// TIA Portal project "Mawomat" (V17) (continued)

               END_IF;

           ELSIF NOT #statSwitchControl OR NOT #statSwitchEnable THEN //if no output enable or switch check then

               IF #statControl THEN

                   #oStatus := 8;

               ELSIF NOT #statControl THEN

                   #oStatus := 2;

               END_IF;

           END_IF;

       ELSE
           #oStatus := 0;

       END_IF;

   END_REGION ;


   REGION Reseting impuls
       // Samokasowanie sygnalow
       #statFaultReset := false;

       IF #inAutoOff THEN

           #statTurnOn := FALSE;

       END_IF;

   END_REGION ;

   REGION Status code


   END_REGION

   REGION Rewriting TO outputs

       #inCmdOper.%X0 := #statManAuto;
       #inCmdOper.%X1 := #statSymOn;
       #inCmdOper.%X2 := #statSwitchEnable;
       #inCmdOper.%X3 := #statManTurnOn;
       #inCmdOper.%X4 := #statManDirection;
       #inCmdOper.%X6 := #statSwitchControl;

       #inCmdOperImp.%X0 := #statFaultReset;

       #oControlMode := #statControlMode;

       #oFault := #statFault;

       #inTurnOn := #statTurnOn;

       #oControl := #statControl;

   END_REGION
END_FUNCTION_BLOCK

// folder: DV

FUNCTION_BLOCK "DV_Objects"   // FB6, LAD
{ S7_Optimized_Access := 'TRUE' }
VERSION : 0.1
   VAR
      dv1 : "DV_Class";
   END_VAR
BEGIN

REGION Network 2 (SCL)
   #dv1();
END_REGION
END_FUNCTION_BLOCK

FUNCTION_BLOCK "DV_Class"   // FB302, SCL
{ S7_Optimized_Access := 'TRUE' }
VERSION : 0.1
   VAR_INPUT
      inActivateObject : Bool := true;   // Aktywowanie działania obiektu
      inTurnOnConfirm : Bool;   // Potwierdzenie załączenia
      inTurnOffConfirm : Bool;   // Potwierdzenie wyłączenia
      inCircBreaker : Bool;   // Gotowość obiektu - rozłącznik
      inPTC : Bool;   // Gotowość obiektu - PTC
      inReadySpare : Bool := true;   // Gotowość obiektu - rezerwa
      inReadySpare2 : Bool := true;   // Gotowość obiektu - rezerwa
      inLocalMode : Bool;   // Tryb lokalny
      inRemoteMode : Bool;   // Tryb remontowy
      inExtFault : Bool;   // Błąd zewnętrzny
      inLockAutoMan : Bool;   // Blokada przełączenia trybu Auto-Manual
      inInterlock : Bool;   // Interlok
      inNoNc : Bool;   // Zawór NO - 1, potw zał - zamkn.; wył-otw
      inGlobalAckFault : Bool;   // Globalny reset
      inAutoOff : Bool;   // Resetowanie sterowania na końcu
      inTurnOnDelay : DInt;   // Czas opóźnienia załączenia [s]
      inTurnOffDelay : DInt;   // Czas opóźnienia wyłączenia [s]
      inAlarmDelay : DInt;   // Czas opóźnienia alarmu od potwierdzeń [s]
   END_VAR
   VAR_OUTPUT
      oControl : Bool;   // Wyjście sterujące
      oAckFault : Bool;   // Wyjście reset obiektu
      oFault : Bool;   // Wyjście awaria
      oFaultCode : Byte;   // Kod awarii
      oStatusCode : Word;   // Kod statusu
      oStatus : Int;   // Status ( 1-awaria; 2-Zamkn; 4-Otwieranie; 8-Otwarte; 16-Zamykanie)
      oControlMode : Int;   // Tryb pracy (1-remont; 2-lokal; 4-manual; 8-auto)
   END_VAR
   VAR_IN_OUT
      inTurnOn : Bool;   // Załączanie z programu
      inCmdOper : Word := 16#5;   // Komendy manualne
      inSimOper : Word;   // Komendy symulacji
      inCmdOperImp : Word;   // Komendy impulsowe
   END_VAR
   VAR
      statReady : Bool;
      statManAuto : Bool;
      statSymOn : Bool;
      statSwitchEnable : Bool;
      statManTurnOn : Bool;
      statManDirection : Bool;
      statSwitchControl : Bool;
      statFaultReset : Bool;
      statActivate : Bool;
      statTurnOn : Bool;
      statTurnOnConfirm : Bool;
      statTurnOffConfirm : Bool;
      statLocal : Bool;
      statRemote : Bool;
      statExtFault : Bool;
      statLockAutoMan : Bool;
      statInterlock : Bool;
      statNoNc : Bool;
      tofTurnOnDelay : TON_TIME;
      tofTurnOffDelay : TOF_TIME;
      tonAlarm : TON_TIME;
      statAlarmStart : Bool;
      statFault : Bool;
      statControlMode : Int;
      statControl : Bool;
      statTmrOnOff : Bool;
      trigGlobalReset : R_TRIG;
   END_VAR
BEGIN
   REGION Activation object - condition to execute function
       IF NOT #inActivateObject THEN
           #inTurnOn := FALSE;
           #inCmdOper := 0;
           #inSimOper := 0;
           #inCmdOperImp := 0;

           #oControl := FALSE;
           #oAckFault := FALSE;
           #oFault := FALSE;
           #oFaultCode := 0;
           #oStatusCode := 0;
           #oStatus := 0;
           #oControlMode := 0;

           RETURN;

       END_IF;

   END_REGION

   REGION Rewriting inputs

       //Operator Control Word
       #statManAuto := #inCmdOper.%X0;
       #statSymOn := #inCmdOper.%X1;
       #statSwitchEnable := #inCmdOper.%X2;
       #statManTurnOn := #inCmdOper.%X3;
       #statManDirection := #inCmdOper.%X4;
       #statSwitchControl := #inCmdOper.%X6;

       //Operator Control Word Impulses
       #trigGlobalReset(CLK:=#inGlobalAckFault);

       #statFaultReset := #trigGlobalReset.Q OR #inCmdOperImp.%X0;

   END_REGION

   REGION Rewriting inputs or simulation signals to statics

       IF NOT #statSymOn THEN

           #statTurnOn := #inTurnOn;
           #statTurnOnConfirm := #inTurnOnConfirm;
           #statTurnOffConfirm := #inTurnOffConfirm;
           #statReady := #inCircBreaker AND #inPTC AND #inReadySpare AND #inReadySpare2 ;
           #statLocal := #inLocalMode;
           #statRemote := #inRemoteMode;
           #statExtFault := #inExtFault;
           #statLockAutoMan := #inLockAutoMan;
           #statInterlock := #inInterlock;
           #statNoNc := #inNoNc;

           //Rewriting inputs to simulation bits when simulotion is to switch fluently
           #inSimOper.%X0 := #statActivate;
           #inSimOper.%X1 := #statTurnOn;
           #inSimOper.%X2 := #statTurnOnConfirm;
           #inSimOper.%X3 := #statTurnOffConfirm;
           #inSimOper.%X4 := #statReady;
           #inSimOper.%X5 := #statLocal;
           #inSimOper.%X6 := #statRemote;
           #inSimOper.%X7 := #statExtFault;
           #inSimOper.%X8 := #statLockAutoMan;
           #inSimOper.%X9 := #statInterlock;
           #inSimOper.%X10 := #statNoNc;

       ELSE

           #statActivate := #inSimOper.%X0;
           #statTurnOn := #inSimOper.%X1;
           #statTurnOnConfirm := #inSimOper.%X2;
           #statTurnOffConfirm := #inSimOper.%X3;
           #statReady:= #inSimOper.%X4;
           #statLocal := #inSimOper.%X5;
           #statRemote := #inSimOper.%X6;
           #statExtFault := #inSimOper.%X7;
           #statLockAutoMan := #inSimOper.%X8;
           #statInterlock := #inSimOper.%X9;
           #statNoNc := #inSimOper.%X10;

       END_IF;


   END_REGION

   REGION Control Mode

       IF #statRemote THEN

           #statControlMode := 1;

       ELSIF #statLocal THEN

           #statControlMode := 2;

       ELSIF NOT #statManAuto AND NOT #statLockAutoMan THEN

           #statControlMode := 4;

       ELSIF #statManAuto AND NOT #statLockAutoMan THEN

           #statControlMode := 8;

       END_IF;

   END_REGION

   REGION TurnOn/Off Delay

       #tofTurnOnDelay(IN := #statTurnOn,
                       PT := 1000 * #inTurnOnDelay);

       #tofTurnOffDelay(IN := #statTurnOn,
                        PT := 1000 * #inTurnOffDelay);

       IF #tofTurnOnDelay.Q THEN

           #statTmrOnOff := TRUE;

       END_IF;

       IF NOT #tofTurnOffDelay.Q THEN

           #statTmrOnOff := FALSE;

       END_IF;
   END_REGION

   REGION Fault 
       //Zerowanie czasu awari przy zmianie sterowanie podczas ruchu - czy to w ogole cokolwiek robi???

       //Alarm from switching control 
       #statAlarmStart :=
       #statSwitchControl AND //is switch controling on
       #statSwitchEnable AND //is objects output is eneble to turn on
       #statControlMode<>2 AND //in local mode there is no alarm
       #statControlMode<>1 AND //in remote mode there is no alarm
       (
       (#statControl XOR #statTurnOnConfirm) OR //xor  0110 - if A and B have different state then =1
       (NOT #statControl XOR #statTurnOffConfirm) OR
       (#statTurnOnConfirm AND #statTurnOffConfirm) OR
       (NOT #statTurnOnConfirm AND NOT #statTurnOffConfirm)
       )
       ;
       //#tonAlarm.PT := DINT_TO_TIME(1000 * #AlarmDelay);
       //Generating switching alarm after delay
       #tonAlarm(IN := #statAlarmStart,
                 PT:=DINT_TO_TIME(1000 * #inAlarmDelay));


       //Generating fault
       IF #tonAlarm.Q OR NOT #statReady OR #statExtFault THEN

           #statFault := TRUE;

       ELSIF #statFaultReset THEN

           #statFault := FALSE;

       END_IF;

       //Fault reset 
       // IF #statFaultReset THEN
       //     #statFault := FALSE;


       // END_IF;

       //Fault code
       #oFaultCode.%X0 := #tonAlarm.Q;
       #oFaultCode.%X1 := NOT #statReady;
       #oFaultCode.%X2 := #statExtFault;
       #oFaultCode.%X3 := NOT #inCircBreaker;
       #oFaultCode.%X4 := NOT #inPTC;
       #oFaultCode.%X5 := NOT #inReadySpare;
       #oFaultCode.%X6 := NOT #inReadySpare2;

   END_REGION

   REGION Command locks

       IF #statControlMode = 8 AND #statLockAutoMan THEN

           #statManAuto := TRUE;

       ELSIF #statControlMode = 4 AND #statLockAutoMan THEN

           #statManAuto := FALSE;

       END_IF;

       // Writing states from Local to Manual when object when switching Local to Manual
       IF #statControlMode = 2 THEN

           #statManAuto := FALSE;

           IF #statTurnOffConfirm THEN

               #statTurnOn := FALSE;

           ELSIF #statTurnOnConfirm THEN

               #statTurnOn := TRUE;

           END_IF;

       END_IF;

       // Writing states from Auto to Manual when object when switching Auto to Manual
       // Przypadek gdy ktos z wlaczonym automatycznie urz. przechodzi na tryb zdalny-reczny
       IF #statControlMode = 8 THEN

           #statManTurnOn := #statTurnOn;
           #statManDirection := #statNoNc;

       END_IF;

       //Resetowanie rozkazu zalaczenia w trybie manualnym po awarii
       IF #statFault THEN

           #statManTurnOn := FALSE;

       END_IF;




   END_REGION

   REGION Control output

       #statControl :=
       #statSwitchEnable AND
       NOT #statInterlock AND
       //NOT #statFault AND - awaria nie powoduje zmiany stanu zaworu
       ((#statControlMode = 8 AND #statTmrOnOff) OR
       (#statControlMode = 4 AND #statManTurnOn));

   END_REGION

   REGION Reset Control

       #oAckFault := #statFaultReset;

   END_REGION ;

   REGION Device status code
       IF #statFault THEN
           #oStatus := 1;

       ELSIF #statControlMode = 1 THEN
           #oStatus := 2;

       ELSIF #statControlMode = 2 THEN

           IF #statTurnOnConfirm THEN

               IF NOT #statNoNc THEN
                   #oStatus := 8;
               ELSE
                   #oStatus := 2;
               END_IF;

           ELSIF #statTurnOffConfirm THEN

               IF NOT #statNoNc THEN
                   #oStatus := 2;
               ELSE
                   #oStatus := 8;
               END_IF;

           ELSIF #statControl THEN

               IF NOT #statNoNc THEN
                   #oStatus := 4;
               ELSE
                   #oStatus := 16;
               END_IF;

           ELSIF NOT #statControl THEN

               IF NOT #statNoNc THEN
                   #oStatus := 16;
               ELSE
                   #oStatus := 4;
               END_IF;
           END_IF;

       ELSIF #statControlMode > 2 THEN

           IF #statSwitchControl AND #statSwitchEnable THEN

               IF #statControl AND NOT #statTurnOffConfirm AND #statTurnOnConfirm THEN

                   IF NOT #statNoNc THEN
                       #oStatus := 8;
                   ELSE
                       #oStatus := 2;
                   END_IF;

               ELSIF NOT #statControl AND NOT #statTurnOnConfirm AND #statTurnOffConfirm THEN

                   IF NOT #statNoNc THEN
                       #oStatus := 2;
                   ELSE
                       #oStatus := 8;
                   END_IF;

               ELSIF #statControl THEN

                   IF NOT #statNoNc THEN
                       #oStatus := 4;
                   ELSE
                       #oStatus := 16;
                   END_IF;

               ELSIF NOT #statControl THEN

                   IF NOT #statNoNc THEN
                       #oStatus := 16;
                   ELSE
                       #oStatus := 4;
                   END_IF;

               END_IF;

           ELSIF NOT #statSwitchControl OR NOT #statSwitchEnable THEN //if no output enable or switch check then

               IF #statControl THEN

                   IF NOT #statNoNc THEN
                       #oStatus := 8;
                   ELSE
                       #oStatus := 2;
                   END_IF;

               ELSIF NOT #statControl THEN

                   IF NOT #statNoNc THEN
                       #oStatus := 2;
                   ELSE
                       #oStatus := 8;
                   END_IF;

               END_IF;

           END_IF;

       ELSE
           #oStatus := 0;

       END_IF;

   END_REGION ;


   REGION Reseting impuls
       // Samokasowanie sygnalow
       #statFaultReset := false;

       IF #inAutoOff THEN

           #statTurnOn := FALSE;

       END_IF;

   END_REGION ;

   REGION Status code


   END_REGION

   REGION Rewriting TO outputs

       #inCmdOper.%X0 := #statManAuto;
       #inCmdOper.%X1 := #statSymOn;
       #inCmdOper.%X2 := #statSwitchEnable;
       #inCmdOper.%X3 := #statManTurnOn;
       #inCmdOper.%X4 := #statManDirection;
       #inCmdOper.%X6 := #statSwitchControl;

       #inCmdOperImp.%X0 := #statFaultReset;

       #oControlMode := #statControlMode;

       #oFault := #statFault;

       #inTurnOn := #statTurnOn;

       #oControl := #statControl;
   END_REGION
END_FUNCTION_BLOCK

// folder: LSim

FUNCTION_BLOCK "LSim_PT1"   // FB50, SCL
{ S7_Optimized_Access := 'TRUE' }
VERSION : 2.01
   VAR_INPUT
      calcParam : Bool;   // recalculate with new parameters
      input : Real;   // input signal
      tmLag1 : Real := 1.0;   // time constant T1 [sec]
      gain : Real := 1.0;   // gain factor
      cycle : Real := 0.1;   // cyclic time [sec]
      maxOut : Real := 100.0;   // max. output limit
      minOut : Real;   // min. output limit
      reset : Bool;   // resets all relevant parameters to ‘0’ including the output
   END_VAR
   VAR_OUTPUT
      error : Bool;   // error (#tmLag1 <= 0)
      status : Word;   // status (if #tmLag1 <= 0 then status = 16#8001)
      maxReached : Bool;   // output has reached max. limit
      minReached : Bool;   // output has reached min. limit
      output : Real;   // output signal (if #error = FALSE)
   END_VAR
   VAR
      statRf1 : Real;
      statRe1 : Real;
      statOverfirst : Bool;
      statOutput : Real;
   END_VAR
BEGIN
   //=============================================================================
   //SIEMENS AG
   //(c)Copyright 2017 All Rights Reserved
   //-----------------------------------------------------------------------------
   //Library:       Library for Controlled System Simulation
   //Tested with:   S7-1500 FW V2.0 / S7-1200 FW V4.2
   //Engineering:   STEP 7 V14 Upd2 (TIA Portal)
   //Restrictions:  Cyclic interrupt
   //Requirements:  memory card needed for S7-1500
   //Functionality: Simulation of a PT1-System
   //
   //              gain
   //  F(p) = ---------------
   //          tmLag1 * p + 1
   //          
   //  Call the simulation in a cyclic interrupt with
   //  cyclic interrupt time at least = tmLag1/10!
   //-----------------------------------------------------------------------------
   //Change log table:
   //Version  Date       Expert in charge                Changes applied
   //02.00.00 03.02.2016 Siemens Industry Online Support Release (STEP 7 V13 SP1)
   //02.00.01 02.03.2017 Siemens Industry Online Support Release (STEP 7 V14)
   //=============================================================================
   // check parameter
   IF #tmLag1 <= 0 THEN
     #error := TRUE;
     #status := W#16#8001;     // Parameter Error
     #statOutput := 0;
     #output := 0;
     RETURN;
   ELSE
     #error := FALSE;
     #status := W#16#0000;     // no error
   END_IF;

   IF #calcParam = True OR NOT #statOverfirst THEN
     #statOverfirst:=1;
   // Z-parameters For Laplace PT1-System
   #statRe1 := - EXP(-#cycle/#tmLag1);
   #statRf1 := #gain*(1 + #statRe1);
   END_IF;

   // Differencial Equation of PT1-System
   #statOutput := #input*#statRf1 - #statOutput*#statRe1;

   // max limit of acutating variable
   IF #statOutput > #maxOut THEN
     #statOutput := #maxOut;
     #maxReached:= True;
   ELSE
     #maxReached := False;
   END_IF;

   // min limit of acutating variable
   IF #statOutput < #minOut THEN
     #statOutput := #minOut;
     #minReached := True;
   ELSE
     #minReached := False;
   END_IF;

   IF #reset THEN
     #statOutput := 0;
   END_IF;

   #output := #statOutput;
END_FUNCTION_BLOCK

FUNCTION_BLOCK "LSim_PT1asym"   // FB51, SCL
{ S7_Optimized_Access := 'TRUE' }
VERSION : 2.01
   VAR_INPUT
      calcParam : Bool;   // recalculate with new parameters
      input : Real;   // input signal
      tmLag1up : Real := 1.0;   // time constant T1 [sec] rising input
      tmLag1down : Real := 10.0;   // time constant T1 [sec] falling input
      gain : Real := 1.0;   // gain factor
      cycle : Real := 0.1;   // cyclic time [sec]
      maxOut : Real := 100.0;   // max. output limit
      minOut : Real;   // min. output limit
      reset : Bool;   // resets all relevant parameters to ‘0’ including the output
   END_VAR
   VAR_OUTPUT
      error : Bool;   // error (#tmLag1 <= 0 or #tmLag2 <= 0)
      status : Word;   // status (if #error = TRUE then status = 16#8001)
      maxReached : Bool;   // output has reached max. limit
      minReached : Bool;   // output has reached min. limit
      output : Real;   // output signal (if #error = FALSE)
   END_VAR
   VAR
      statRxn1 : Real;   // delayed input signal (n-1)
      statRyn1 : Real;   // delayed output signal (n-1)
      statRf1up : Real;   // Z-parameter 1 (rising xn)
      statRe1up : Real;   // Z-parameter 2 (rising xn)
      statRf1dn : Real;   // Z-parameter 1 (falling xn)
      statRe1dn : Real;   // Z-parameter 2 (falling xn)
      statRf1 : Real;   // active Z-parameter 1
      statRe1 : Real;   // active Z-parameter 2
      statOverfirst : Bool;
      statOutput : Real;
   END_VAR
BEGIN
   //=============================================================================
   //SIEMENS AG
   //(c)Copyright 2017 All Rights Reserved
   //-----------------------------------------------------------------------------
   //Library:       Library for Controlled System Simulation
   //Tested with:   S7-1500 FW V2.0 / S7-1200 FW V4.2
   //Engineering:   STEP 7 V14 Upd2 (TIA Portal)
   //Restrictions:  Cyclic interrupt
   //Requirements:  memory card needed for S7-1500
   //Functionality: Simulation of a PT1-System with two different Time-Constants
   //
   //  tmLag1up: Time-Constant for positive Inputsignal changes 
   //  tmLag1down: Time-Constant for negative Inputsignal changes
   //  
   //                gain
   //  Fup(p) = ----------------
   //           tmLag1up * p + 1
   //          
   //                    gain
   //  Fdown(p) = ------------------
   //             tmLag1down * p + 1
   //          
   //  Call the simulation in a cyclic interrupt with
   //  //  cyclic interrupt time at least = tmLag1/10!
   //-----------------------------------------------------------------------------
   //Change log table:
   //Version  Date       Expert in charge                Changes applied
   //02.00.00 03.02.2016 Siemens Industry Online Support Release (STEP 7 V13 SP1)
   //02.00.01 02.03.2017 Siemens Industry Online Support Release (STEP 7 V14)
   //=============================================================================

   // check parameter
   IF #tmLag1up <= 0 OR #tmLag1down <= 0 THEN
     #error := TRUE;
     #status := W#16#8001;     // Parameter Error
     #statOutput := 0;
     #output := 0;
     RETURN;
   ELSE
     #error := FALSE;
     #status := W#16#0000;     // no error
   END_IF;

   IF #calcParam = True OR NOT #statOverfirst THEN
     #statOverfirst:=1;
   // Z-parameters for Laplace PT1-System (rising signal change)
   #statRe1up := - EXP(-#cycle/#tmLag1up);
   #statRf1up := #gain*(1 + #statRe1up);
   // Z-parameters for Laplace PT1-System (falling signal change)
   #statRe1dn := - EXP(-#cycle/#tmLag1down);
   #statRf1dn := #gain*(1 + #statRe1dn);
   END_IF;

   // save delayed output signals
   #statRyn1:= #statOutput;

   // Change the parameter sets, dependent to Input Change
   IF (#input - #statRxn1) > 0 THEN
     #statRf1 := #statRf1up;
     #statRe1 := #statRe1up;
   ELSIF (#input - #statRxn1) < 0 THEN
      #statRf1 := #statRf1dn;
      #statRe1 := #statRe1dn;
   ELSE
     ;
   END_IF;

   // Differencial Equation of PT1-System
   #statOutput := #input*#statRf1 - #statRyn1*#statRe1;

   // save delayed input signals
   #statRxn1 := #input;

   // max limit of acutating variable
   IF #statOutput > #maxOut THEN
     #statOutput := #maxOut;
     #maxReached:= True;
   ELSE
     #maxReached := False;
   END_IF;

   // min limit of acutating variable
   IF #statOutput < #minOut THEN
     #statOutput := #minOut;
     #minReached := True;
   ELSE
     #minReached := False;
   END_IF;

   IF #reset THEN
     #statOutput := 0;
   END_IF;

   #output := #statOutput;
END_FUNCTION_BLOCK

FUNCTION_BLOCK "LSim_PT2osc"   // FB52, SCL
{ S7_Optimized_Access := 'TRUE' }
VERSION : 2.01
   VAR_INPUT
      calcParam : Bool;   // recalculate with new parameters
      input : Real;   // input signal
      omega : Real := 2.0;   // angular frequency of the undampened vibrations [1/sec]
      damp : Real := 0.2;   // damping (0 < D < 1)
      gain : Real := 1.0;   // gain factor
      cycle : Real := 0.1;   // cyclic time [sec]
      maxOut : Real := 100.0;   // max. output limit
      minOut : Real;   // min. output limit
      reset : Bool;   // resets all relevant parameters to ‘0’ including the output
   END_VAR
   VAR_OUTPUT
      error : Bool;   // error (0 >= damp >= 1 or #omega <= 0)
      status : Word;   // status (if #error = TRUE then status = 16#8001)
      maxReached : Bool;   // output has reached max. limit
      minReached : Bool;   // output has reached min. limit
      output : Real;   // output signal (if #error = FALSE)
   END_VAR
   VAR
      statRxn2 : Real;   // delayed input signal (n-2)
      statRxn1 : Real;   // delayed input signal (n-1)
      statRyn2 : Real;   // delayed output signal (n-2)
      statRyn1 : Real;   // delayed output signal (n-1)
      statRb1 : Real;
      statRb2 : Real;
      statRa1 : Real;
      statRa2 : Real;
      statRo : Real;
      statSigma : Real;
      statNue : Real;
      statOverfirst : Bool;
      statOutput : Real;
   END_VAR
BEGIN
   //=============================================================================
   //SIEMENS AG
   //(c)Copyright 2017 All Rights Reserved
   //-----------------------------------------------------------------------------
   //Library:       Library for Controlled System Simulation
   //Tested with:   S7-1500 FW V2.0 / S7-1200 FW V4.2
   //Engineering:   STEP 7 V14 Upd2 (TIA Portal)
   //Restrictions:  Cyclic interrupt
   //Requirements:  memory card needed for S7-1500
   //Functionality: Simulation of a vibrating PT2-System
   //
   //                  gain
   //  F(p) = ----------------------------------
   //         SQR(p/omega) + 2*damp*p/omega + 1
   //          
   //  Call the simulation in a cyclic interrupt with
   //  cyclic interrupt time at least = tmLag1/10!
   //-----------------------------------------------------------------------------
   //Change log table:
   //Version  Date       Expert in charge                Changes applied
   //02.00.00 03.02.2016 Siemens Industry Online Support Release (STEP 7 V13 SP1)
   //02.00.01 02.03.2017 Siemens Industry Online Support Release (STEP 7 V14)
   //=============================================================================

   // check parameter
   IF #damp >= 1 OR #damp <= 0 OR #omega <= 0 THEN
     #error := TRUE;
     #status := W#16#8001;
     #statRxn1 := 0.0;
     #statRyn1 := 0.0;
     #statRxn2 := 0.0;
     #statRyn2 := 0.0;
     #statOutput := 0;
     #output := 0;
     RETURN;
   ELSE
     #error := FALSE;
     #status := W#16#0000;     // no error 
   END_IF;

   // calculates the z-parameter for the difference equatation
   IF #calcParam = True THEN
   // Calculate z-parameters for oscillating PT2-System
   #statRo := EXP(-2*#omega*#damp*#cycle);
   #statSigma := (COS(#omega * #cycle * SQRT(1 - SQR(#damp)))) * EXP(-#damp*#omega*#cycle);
   #statNue := (SIN(#omega*#cycle*SQRT(1-SQR(#damp)))) * (EXP(-#damp*#omega*#cycle)) * (#damp / SQRT(1 - SQR(#damp)));
   #statRa1 := -2*#statSigma;
   #statRa2 := #statRo;
   #statRb1 := #gain*(1 - #statSigma - #statNue);
   #statRb2 := #gain*(#statRo - #statSigma + #statNue);
   END_IF;

   // reset Memory
   IF #reset = True THEN
     #statRxn1 := 0.0;
     #statRyn1 := 0.0;
     #statRxn2 := 0.0;
     #statRyn2 := 0.0;
     #statOutput:=0;
     #error := False;
     #status := W#16#0000;
   END_IF;

   // save delayed output signals
   #statRyn2:=#statRyn1;
   #statRyn1:= #statOutput;

   // difference equatation for PT2-System
   #statOutput := #statRxn1* #statRb1 + #statRxn2*#statRb2 - #statRyn1*#statRa1 - #statRyn2*#statRa2;

   // save delayed input signals
   #statRxn2 := #statRxn1;
   #statRxn1 := #input;

   // max limit of acutating variable
   IF #statOutput > #maxOut THEN
     #statOutput := #maxOut;
     #maxReached:= True;
   ELSE
     #maxReached := False;
   END_IF;

   // min limit of acutating variable
   IF #statOutput < #minOut THEN
     #statOutput := #minOut;
     #minReached := True;
   ELSE
     #minReached := False;
   END_IF;

   #output := #statOutput;
END_FUNCTION_BLOCK

FUNCTION_BLOCK "LSim_PT2aper"   // FB53, SCL
{ S7_Optimized_Access := 'TRUE' }
VERSION : 2.01
   VAR_INPUT
      calcParam : Bool;   // recalculate with new parameters
      input : Real;   // input signal
      tmLag1 : Real := 2.0;   // time constant T1 [sec]
      tmLag2 : Real := 0.2;   // time constant T2 [sec]
      gain : Real := 1.0;   // gain factor
      cycle : Real := 0.1;   // cyclic time [sec]
      maxOut : Real := 100.0;   // max. output limit
      minOut : Real;   // min. output limit
      reset : Bool;   // resets all relevant parameters to ‘0’ including the output
   END_VAR
   VAR_OUTPUT
      error : Bool;   // error (#tmLag1 <= 0 or #tmLag2 <= 0 or #tmLag1 = #tmLag2)
      status : Word;   // status (if #error = TRUE then status = 16#8001)
      maxReached : Bool;   // output has reached max. limit
      minReached : Bool;   // output has reached min. limit
      output : Real;   // output signal (if #error = FALSE)
   END_VAR
   VAR
      statRxn2 : Real;   // delayed input signal (n-2)
      statRxn1 : Real;   // delayed input signal (n-1)
      statRyn2 : Real;   // delayed output signal (n-2)
      statRyn1 : Real;   // delayed output signal (n-1)
      statRf1 : Real;
      statRf2 : Real;
      statRe1 : Real;
      statRe2 : Real;
      statAlpha : Real;
      statBeta : Real;
      statGamma : Real;
      statDelta : Real;
      statOverfirst : Bool;
      statOutput : Real;   // Output signal
   END_VAR
BEGIN
   //=============================================================================
   //SIEMENS AG
   //(c)Copyright 2017 All Rights Reserved
   //-----------------------------------------------------------------------------
   //Library:       Library for Controlled System Simulation
   //Tested with:   S7-1500 FW V2.0 / S7-1200 FW V4.2
   //Engineering:   STEP 7 V14 Upd2 (TIA Portal)
   //Restrictions:  Cyclic interrupt
   //Requirements:  memory card needed for S7-1500
   //Functionality: Simulation of a aperiodic PT2-System
   //  
   //                    gain
   //  F(p) = -----------------------------
   //         (tmLag1*p + 1)*(tmLag2*p + 1)
   //         
   //  Call the simulation in a cyclic interrupt with
   //  cyclic interrupt time at least = tmLag1/10!
   //-----------------------------------------------------------------------------
   //Change log table:
   //Version  Date       Expert in charge                Changes applied
   //02.00.00 03.02.2016 Siemens Industry Online Support Release (STEP 7 V13 SP1)
   //02.00.01 02.03.2017 Siemens Industry Online Support Release (STEP 7 V14)
   //=============================================================================

   // check parameter
   IF #tmLag1 <= 0 OR #tmLag2 <= 0 OR #tmLag1 = #tmLag2 THEN
     #error := TRUE;
     #status := W#16#8001;     // Parameter Error
     #statRxn1 := 0.0;
     #statRyn1 := 0.0;
     #statRxn2 := 0.0;
     #statRyn2 := 0.0;
     #statOutput := 0;
     #output := 0;
     RETURN;
   ELSE
     #error := FALSE;
     #status := W#16#0000;     // no error
   END_IF;

   // calculates the z-parameter for the difference equatation
   IF #calcParam = True OR NOT #statOverfirst THEN
     #statOverfirst := 1;
     // Calculate z-parameters for IT1-System
     #statAlpha := EXP(- #cycle / #tmLag1);
     #statBeta := EXP(- #cycle / #tmLag2);
     #statGamma := #tmLag1 / (#tmLag1 - #tmLag2);
     #statDelta := #tmLag2 / (#tmLag1 - #tmLag2);
     #statRe1 := - #statAlpha - #statBeta;
     #statRe2 := #statAlpha * #statBeta;
     #statRf1 := #gain * (1 - #statGamma * #statAlpha + #statDelta * #statBeta);
     #statRf2 := #gain * (#statAlpha * #statBeta - #statGamma * #statBeta + #statAlpha * #statDelta);
   END_IF;

   // reset Memory
   IF #reset = True THEN
     #statRxn1 := 0.0;
     #statRyn1 := 0.0;
     #statRxn2 := 0.0;
     #statRyn2 := 0.0;
     #statOutput := 0;
   END_IF;
   //save delayed input signals
   #statRxn2 := #statRxn1;
   #statRxn1 := #input;

   //save delayed output signals
   #statRyn2:=#statRyn1;
   #statRyn1:= #statOutput;

   // difference equatation of the PT2-System
   #statOutput := #statRxn1* #statRf1 + #statRxn2*#statRf2 - #statRyn1*#statRe1 - #statRyn2*#statRe2;

   // max limit of acutating variable
   IF #statOutput > #maxOut THEN
     #statOutput := #maxOut;
     #maxReached:= True;
   ELSE
     #maxReached := False;
   END_IF;

   // min limit of acutating variable
   IF #statOutput < #minOut THEN
     #statOutput := #minOut;
     #minReached := True;
   ELSE
     #minReached := False;
   END_IF;

   #output := #statOutput;
END_FUNCTION_BLOCK

FUNCTION_BLOCK "LSim_PT3"   // FB54, SCL
{ S7_Optimized_Access := 'TRUE' }
VERSION : 2.01
   VAR_INPUT
      input : Real;   // input variable
      tmLag1 : Real := 29.0;   // time lag 1 in s
      tmLag2 : Real := 17.5;   // time lag 2 in s
      tmLag3 : Real := 3.1;   // time lag 3 in s
      gain : Real := 1.0;   // proportional gain
      disturb : Real;   // disturbance variable (additional to "input")
      cycle : Real := 0.1;   // sample time [in sec]
      reset : Bool;   // complete restart (#output = #input)
   END_VAR
   VAR_OUTPUT
      error : Bool;   // error (#tmLag1 <= 0 or #tmLag2 <= 0 or #tmLag3 <= 0)
      status : Word;   // status (if #error = TRUE then status = 16#8001)
      output : Real;   // output signal (if #error = FALSE)
   END_VAR
   VAR
      statFback1 : Real;   // feedback path value 1
      statFback2 : Real;   // feedback path value 2
      statFback3 : Real;   // feedback path value 3
   END_VAR
   VAR_TEMP
      tempHvar : Real;   // help variable
      tempCycleR : Real;   // cycle to real
      tempTmLag1R : Real;   // time lag 1 to real
      tempTmLag2R : Real;   // time lag 2 to real
      tempTmLag3R : Real;   // time lag 3 to real
      tempOutvNew : Real;   // new output variable
   END_VAR
BEGIN
   //=============================================================================
   //SIEMENS AG
   //(c)Copyright 2017 All Rights Reserved
   //-----------------------------------------------------------------------------
   //Library:       Library for Controlled System Simulation
   //Tested with:   S7-1500 FW V2.0 / S7-1200 FW V4.2
   //Engineering:   STEP 7 V14 Upd2 (TIA Portal)
   //Restrictions:  Cyclic interrupt
   //Requirements:  memory card needed for S7-1500
   //Functionality: Simulation of an PT3-system
   //
   //                               gain
   //  F(p) = ------------------------------------------------------
   //         (tmLag1 * p + 1) * (tmLag2 * p + 1) * (tmLag3 * p + 1)
   //          
   //  Call the simulation in a cyclic interrupt with
   //  cyclic interrupt time at least = tmLag1/10!
   //-----------------------------------------------------------------------------
   //Change log table:
   //Version  Date       Expert in charge                Changes applied
   //02.00.00 03.02.2016 Siemens Industry Online Support Release (STEP 7 V13 SP1)
   //02.00.01 02.03.2017 Siemens Industry Online Support Release (STEP 7 V14)
   //=============================================================================
   // check parameter
   IF #tmLag1 <= 0 OR #tmLag2 <= 0 OR #tmLag3 <= 0 THEN
     #error := TRUE;
     #status := W#16#8001;     // Parameter Error
     #output := #input; //write output data
     #statFback1 := #input; //write static data
     #statFback2 := #input;
     #statFback3 := #input;
     RETURN;
   ELSE
     #error := FALSE;
     #status := W#16#0000;     // no error
   END_IF;

   IF #reset THEN //complete restart routine

     #output := #input;//write output data
     #statFback1 := #input;//write static data
     #statFback2 := #input;
     #statFback3 := #input;

   ELSE //cycle mode routine

     #tempCycleR  := #cycle*1000; //transform data type
     #tempTmLag1R := #tmLag1*1000;
     #tempTmLag2R := #tmLag2*1000;
     #tempTmLag3R := #tmLag3*1000;

     IF #tempCycleR * 0.5 > #tempTmLag1R THEN //limit TM_LAG1
       #tempTmLag1R := #tempCycleR * 0.5;
     END_IF;

     IF #tempCycleR * 0.5 > #tempTmLag2R THEN //limit TM_LAG2
       #tempTmLag2R := #tempCycleR * 0.5;
     END_IF;

     IF #tempCycleR * 0.5 > #tempTmLag3R THEN //limit TM_LAG2
       #tempTmLag3R := #tempCycleR * 0.5;
     END_IF;

     //1. first order lag algorithm
     #tempHvar     := #tempCycleR / (#tempTmLag1R * 2.0); 
     #tempHvar     := (#gain * (#input + #disturb) - #statFback1) * #tempHvar / (#tempHvar + 1.0);
     #tempOutvNew  := #tempHvar + #statFback1;
     #statFback1  := #tempHvar * 2.0 + #statFback1;

     //2. first order lag algorithm
     #tempHvar     := #tempCycleR / (#tempTmLag2R * 2.0); 
     #tempHvar     := ((#tempOutvNew - #statFback2) * #tempHvar) / (#tempHvar + 1.0);
     #tempOutvNew  := #tempHvar + #statFback2;
     #statFback2  := #tempHvar * 2.0 + #statFback2;

     //3. first order lag algorithm
     #tempHvar     := #tempCycleR / (#tempTmLag3R * 2.0); 
     #tempHvar     := ((#tempOutvNew - #statFback3) * #tempHvar) / (#tempHvar + 1.0);
     #tempOutvNew  := #tempHvar + #statFback3;
     #statFback3  := #tempHvar * 2.0 + #statFback3;

     #output := #tempOutvNew; //write output

   END_IF;
END_FUNCTION_BLOCK

FUNCTION_BLOCK "LSim_PDT1"   // FB55, SCL
{ S7_Optimized_Access := 'TRUE' }
VERSION : 2.01
   VAR_INPUT
      calcParam : Bool;   // recalculate with new parameters
      input : Real;   // input signal
      tmLag1 : Real := 2.0;   // time constant T1 [sec]
      tmLag2 : Real := 0.2;   // time constant T2 [sec]
      gain : Real := 1.0;   // gain factor
      cycle : Real := 0.1;   // cyclic time [sec]
      maxOut : Real := 100.0;   // max. output limit
      minOut : Real;   // min. output limit
      reset : Bool;   // resets all relevant parameters to ‘0’ including the output
   END_VAR
   VAR_OUTPUT
      error : Bool;   // error (#tmLag1 <= 0 or #tmLag2 <= 0)
      status : Word;   // status (if #error = TRUE then status = 16#8001)
      maxReached : Bool;   // output has reached max. limit
      minReached : Bool;   // output has reached min. limit
      output : Real;   // output signal (if #error = FALSE)
   END_VAR
   VAR
      statRxn2 : Real;   // delayed input signal (n-2)
      statRxn1 : Real;   // delayed input signal (n-1)
      statRyn2 : Real;   // delayed output signal (n-2)
      statRyn1 : Real;   // delayed output signal (n-1)
      statRb1 : Real;
      statRb0 : Real;
      statRa1 : Real;
      statOverfirst : Bool;
      statOutput : Real;
   END_VAR
BEGIN
   //=============================================================================
   //SIEMENS AG
   //(c)Copyright 2017 All Rights Reserved
   //-----------------------------------------------------------------------------
   //Library:       Library for Controlled System Simulation
   //Tested with:   S7-1500 FW V2.0 / S7-1200 FW V4.2
   //Engineering:   STEP 7 V14 Upd2 (TIA Portal)
   //Restrictions:  Cyclic interrupt
   //Requirements:  memory card needed for S7-1500
   //Functionality: Simulation of an PD-T1 System
   //
   //         gain * (1 + tmLag2*p)
   //  F(p) = ------------------------------
   //            (1 + tmLag1*p)
   //          
   //  Call the simulation in a cyclic interrupt with
   //  cyclic interrupt time at least = tmLag1/10!
   //-----------------------------------------------------------------------------
   //Change log table:
   //Version  Date       Expert in charge                Changes applied
   //02.00.00 03.02.2016 Siemens Industry Online Support Release (STEP 7 V13 SP1)
   //02.00.01 02.03.2017 Siemens Industry Online Support Release (STEP 7 V14)
   //=============================================================================

   // check parameter
   IF #tmLag1 <= 0 OR #tmLag2 <= 0 THEN
     #error := True;
     #status := W#16#8001;     // Parameter Error
     #statRxn1 := 0.0;
     #statRyn1 := 0.0;
     #statRxn2 := 0.0;
     #statRyn2 := 0.0;
     #statOutput := 0;
     #output := 0;
     RETURN;
   ELSE
     #error := FALSE;
     #status := W#16#0000;     // no error
   END_IF;

   // calculates the z-parameter for the difference equatation
   IF #calcParam = True OR NOT #statOverfirst THEN
     #statOverfirst := 1;
   // Calculate z-parameters for oscilating PT2-System
   #statRa1 := -EXP(-#cycle/#tmLag1);
   #statRb0 := #gain *(#tmLag2/#tmLag1);
   #statRb1 := #gain *(1 + #statRa1 - (#tmLag2/#tmLag1));
   END_IF;

   // reset Memory
   IF #reset = True THEN
     #statRxn1 := 0.0;
     #statRyn1 := 0.0;
     #statRxn2 := 0.0;
     #statRyn2 := 0.0;
     #statOutput:=0;
     #error := False;
     #status := W#16#0000;
   END_IF;

   // save delayed output-signals
   #statRyn1:= #statOutput;

   // difference equatation for PT2-system
   #statOutput := #input * #statRb0 +  #statRxn1* #statRb1 - #statRyn1*#statRa1;

   // save delayed input-signals
   #statRxn1 := #input;

   // max limit of acutating variable
   IF #statOutput > #maxOut THEN
     #statOutput := #maxOut;
     #maxReached:= True;
   ELSE
     #maxReached := False;
   END_IF;

   // min limit of acutating variable
   IF #statOutput < #minOut THEN
     #statOutput := #minOut;
     #minReached := True;
   ELSE
     #minReached := False;
   END_IF;

   #output := #statOutput;
END_FUNCTION_BLOCK

FUNCTION_BLOCK "LSim_I"   // FB56, SCL
{ S7_Optimized_Access := 'TRUE' }
VERSION : 2.01
   VAR_INPUT
      calcParam : Bool;   // recalculate with new parameters
      input : Real;   // input signal
      tmLag1 : Real := 1.0;   // time constant T1 [sec]
      cycle : Real := 0.1;   // cyclic time [sec]
      maxOut : Real := 100.0;   // max. output limit
      minOut : Real;   // min. output limit
      reset : Bool;   // resets all relevant parameters to ‘0’ including the output
   END_VAR
   VAR_OUTPUT
      error : Bool;   // error (#tmLag1 <= 0)
      status : Word;   // status (if #tmLag1 <= 0 then status = 16#8001)
      maxReached : Bool;   // output has reached max. limit
      minReached : Bool;   // output has reached min. limit
      output : Real;   // output signal (if #error = FALSE)
   END_VAR
   VAR
      statRxn1 : Real;   // delayed input signal (n-1)
      statRyn1 : Real;   // delayed output signal (n-1)
      statRa1 : Real;
      statRb1 : Real;
      statOverfirst : Bool;
      statOutput : Real;   // output signal
   END_VAR
BEGIN
   //=============================================================================
   //SIEMENS AG
   //(c)Copyright 2017 All Rights Reserved
   //-----------------------------------------------------------------------------
   //Library:       Library for Controlled System Simulation
   //Tested with:   S7-1500 FW V2.0 / S7-1200 FW V4.2
   //Engineering:   STEP 7 V14 Upd2 (TIA Portal)
   //Restrictions:  Cyclic interrupt
   //Requirements:  memory card needed for S7-1500
   //Functionality: Simulation of a I-System
   //
   //             1
   //  F(p) = -----------
   //         (tmLag1*p)
   //          
   //  Call the simulation in a cyclic interrupt with
   //  cyclic interrupt time at least = tmLag1/10!
   //-----------------------------------------------------------------------------
   //Change log table:
   //Version  Date       Expert in charge                Changes applied
   //02.00.00 03.02.2016 Siemens Industry Online Support Release (STEP 7 V13 SP1)
   //02.00.01 02.03.2017 Siemens Industry Online Support Release (STEP 7 V14)
   //=============================================================================

   // check parameter
   IF #tmLag1 <= 0 THEN
     #error := True;
     #status := W#16#8001;     // Parameter Error
     #statRxn1 := 0.0;
     #statRyn1 := 0.0;
     #statOutput := 0;
     #output := 0;
     RETURN;
   ELSE
     #error := FALSE;
     #status := W#16#0000;     // no error
   END_IF;

   // calculates the z-parameter for the difference equatation
   IF #calcParam = True OR NOT #statOverfirst THEN
   #statOverfirst:=1;
     // Calculate z-parameters for IT1-System
   #statRb1 := #cycle/#tmLag1;
   #statRa1 := -1;

   END_IF;

   // reset Memory
   IF #reset = True THEN
     #statRxn1 := 0.0;
     #statRyn1 := 0.0;
     #statOutput:=0;
   END_IF;

   // save delayed output-signals
   #statRyn1:= #statOutput;

   // difference equatation for the I-system
   #statOutput := #statRxn1* #statRb1 - #statRyn1*#statRa1;

   // save delayed input-signals
   #statRxn1 := #input;

   // max limit of acutating variable
   IF #statOutput > #maxOut THEN
     #statOutput := #maxOut;
     #maxReached:= True;
   ELSE
     #maxReached := False;
   END_IF;

   // min limit of acutating variable
   IF #statOutput < #minOut THEN
     #statOutput := #minOut;
     #minReached := True;
   ELSE
     #minReached := False;
   END_IF;

   #output := #statOutput;
END_FUNCTION_BLOCK

FUNCTION_BLOCK "LSim_IT1"   // FB57, SCL
{ S7_Optimized_Access := 'TRUE' }
VERSION : 2.01
   VAR_INPUT
      calcParam : Bool;   // recalculate with new parameters
      input : Real;   // input signal
      tmLag1 : Real := 5.0;   // time constant T1 [sec]
      gain : Real := 1.0;   // gain factor
      cycle : Real := 0.1;   // cyclic time [sec]
      maxOut : Real := 100.0;   // max. output limit
      minOut : Real;   // min. output limit
      reset : Bool;   // resets all relevant parameters to ‘0’ including the output
   END_VAR
   VAR_OUTPUT
      error : Bool;   // error (#tmLag1 <= 0)
      status : Word;   // status (if #tmLag1 <= 0 then status = 16#8001)
      maxReached : Bool;   // output has reached max. limit
      minReached : Bool;   // output has reached min. limit
      output : Real;   // output signal (if #error = FALSE)
   END_VAR
   VAR
      statRxn2 : Real;   // delayed input signal (n-2)
      statRxn1 : Real;   // delayed input signal (n-1)
      statRyn2 : Real;   // delayed output signal (n-2)
      statRyn1 : Real;   // delayed output signal (n-1)
      statRf1 : Real;
      statRf2 : Real;
      statRe1 : Real;
      statRe2 : Real;
      statAlpha : Real;
      statOverfirst : Bool;
      statOutput : Real;   // output signal
   END_VAR
BEGIN
   //=============================================================================
   //SIEMENS AG
   //(c)Copyright 2017 All Rights Reserved
   //-----------------------------------------------------------------------------
   //Library:       Library for Controlled System Simulation
   //Tested with:   S7-1500 FW V2.0 / S7-1200 FW V4.2
   //Engineering:   STEP 7 V14 Upd2 (TIA Portal)
   //Restrictions:  Cyclic interrupt
   //Requirements:  memory card needed for S7-1500
   //Functionality: Simulation of a IT1-System
   //  
   //               gain
   //  F(p) = ------------------
   //         p * (tmLag1*p + 1)
   //         
   //  Call the simulation in a cyclic interrupt with
   //  cyclic interrupt time at least = tmLag1/10!
   //-----------------------------------------------------------------------------
   //Change log table:
   //Version  Date       Expert in charge                Changes applied
   //02.00.00 03.02.2016 Siemens Industry Online Support Release (STEP 7 V13 SP1)
   //02.00.01 02.03.2017 Siemens Industry Online Support Release (STEP 7 V14)
   //=============================================================================


   // check parameter
   IF #tmLag1 <= 0 THEN
     #error := True;
     #status := W#16#8001;     // Parameter Error
     #statRxn1 := 0.0;
     #statRyn1 := 0.0;
     #statRxn2 := 0.0;
     #statRyn2 := 0.0;
     #statOutput := 0;
     #output := 0;
     RETURN;
   ELSE
     #error := FALSE;
     #status := W#16#0000;     // no error
   END_IF;

   // calculates the z-parameter for the difference equatation
   IF #calcParam = True OR NOT #statOverfirst THEN
     #statOverfirst:=1;
   // calculates the z-parameter for the difference equatation of the IT1-System
   #statAlpha := EXP(-#cycle/#tmLag1);
   #statRe1 := -1 - #statAlpha;
   #statRe2 := #statAlpha;
   #statRf1 := #gain*(#cycle +(#statAlpha - 1)*#tmLag1);
   #statRf2 := #gain*(-#statAlpha*#cycle+(1-#statAlpha)*#tmLag1);
   END_IF;

   // reset Memory
   IF #reset = True THEN
     #statRxn1 := 0.0;
     #statRyn1 := 0.0;
     #statRxn2 := 0.0;
     #statRyn2 := 0.0;
     #statOutput:=0;
   END_IF;

   // save delayed output-signals
   #statRyn2:=#statRyn1;
   #statRyn1:= #statOutput;

   // difference equatation for IT1-System
   #statOutput := #statRxn1* #statRf1 + #statRxn2*#statRf2 - #statRyn1*#statRe1 - #statRyn2*#statRe2;

   // save delayed input-signals
   #statRxn2 := #statRxn1;
   #statRxn1 := #input;

   // max limit of acutating variable
   IF #statOutput > #maxOut THEN
   #statOutput := #maxOut;
   #maxReached := True;
   ELSE
     #maxReached := False;
   END_IF;

   // min limit of acutating variable
   IF #statOutput < #minOut THEN
     #statOutput := #minOut;
     #minReached := True;
   ELSE
     #minReached := False;
   END_IF;

   #output := #statOutput;
END_FUNCTION_BLOCK

FUNCTION_BLOCK "LSim_TempProcess"   // FB58, SCL
{ S7_Optimized_Access := 'TRUE' }
VERSION : 2.01
   VAR_INPUT
      inTemp : Real;   // Temperature Input [K] ("useHeatPow" must be FALSE to use this input)
      useHeatPow : Bool := TRUE;   // Use "heatPow" as input
      activHeatPow : Bool;   // Turn on heating ("useHeatPow" must be TRUE to use this input)
      activCoolRth : Bool;   // Turn on cooling by "statRThCool"
      activCoolPow : Bool;   // Turn on cooling by "coolPow"
      coolPow : Real;   // Positive value of energy reduction caused by succeding process [W]
      ambTemp : Real := 20.0;   // Ambient Temperature in °C
      cycle : Real := 0.1;   // Call cycle time in s
      reset : Bool;   // Reset internal variables
   END_VAR
   VAR_OUTPUT
      outTemp : Real;   // [°C]
      interTemp : Real;   // [°C]
   END_VAR
   VAR_IN_OUT
      heatPow : Real;   // Heater Energy in [W]
   END_VAR
   VAR
      statRthTrans1 : Real := 1.5;   // Input thermal resistance in transition to capacitor 1 [K/W]
      statRth1 : Real := 1.0;   // Thermal resistance parallel to thermal capacity 1 [K/W]
      statRthTrans2 : Real := 1.5;   // Thermal resistance for energy transition from capacity 1 to capacity 2 [K/W]
      statRth2 : Real := 1.0;   // Thermal resistance parallel to thermal capacity 2 [K/W]
      statRthCool : Real := 2.0;   // Thermal resistance of cooling device [K/W]
      statCth1 : Real := 10.0;   // Thermal Capacity 1 [Ws/K]
      statCth2 : Real := 30.0;   // Thermal Capacity 2 [Ws/K]
      statZInt1 : Real;   // internal
      statZInt2 : Real;   // internal
      statUc1 : Real;   // internal
      statUc2 : Real;   // internal
      statIth2 : Real;   // internal
   END_VAR
   VAR_TEMP
      tempSumPoint1 : Real;
      tempSumPoint2 : Real;
   END_VAR
BEGIN
   //=============================================================================
   //SIEMENS AG
   //(c)Copyright 2017 All Rights Reserved
   //-----------------------------------------------------------------------------
   //Library:       Library for Controlled System Simulation
   //Tested with:   S7-1500 FW V2.0 / S7-1200 FW V4.2
   //Engineering:   STEP 7 V14 Upd2 (TIA Portal)
   //Restrictions:  Cyclic interrupt
   //Requirements:  memory card needed for S7-1500
   //Functionality: Simulates of an asymmetrical temperature process which can be
   //actively heated and cooled down (also passively).
   //-----------------------------------------------------------------------------
   //Change log table:
   //Version  Date       Expert in charge                Changes applied
   //02.00.00 03.02.2016 Siemens Industry Online Support Release (STEP 7 V13 SP1)
   //02.00.01 02.03.2017 Siemens Industry Online Support Release (STEP 7 V14)
   //=============================================================================
   IF #reset = TRUE THEN
     // Reset all variables
     #statUc1 := 0;
     #statUc2 := 0;
     #statIth2 := 0;
     #tempSumPoint1 := 0;
     #tempSumPoint2 := 0;
     #statZInt1 := 0;
     #statZInt2 := 0;
   END_IF;

   IF #useHeatPow = FALSE THEN
     // Temperature Input will be used, so "heatPow" will be used as output
     #heatPow := ((#inTemp - #ambTemp - #statUc1) / #statRthTrans1);
   END_IF;

   // Calculate fist summing point
   IF (#activHeatPow = TRUE) OR (#useHeatPow = FALSE) THEN
     #tempSumPoint1 := #heatPow - (#statUc1 / #statRth1) - #statIth2;
   ELSE
     #tempSumPoint1 := 0 - (#statUc1 / #statRth1) - #statIth2;
   END_IF;

   // Calculate integrator 1
   #statUc1 := #statUc1 + (((#tempSumPoint1 / #statCth1) + #statZInt1) * #cycle * 0.5);
   #statZInt1 := #tempSumPoint1 / #statCth1;

   // Calculate intermidiate temperature
   #interTemp := #statUc1 + #ambTemp;

   // Calculate thermal power flow from Integrator 1 to Integrator 2
   #statIth2 := ((#statUc1 - #statUc2) / #statRthTrans2);

   // Calculate summing point 2
   IF #activCoolPow = TRUE THEN
     #tempSumPoint2 := #statIth2 - (#statUc2 / #statRth2) - #coolPow;
   ELSE
     #tempSumPoint2 := #statIth2 - (#statUc2 / #statRth2);
   END_IF;

   IF #activCoolRth = TRUE THEN
     // Cooling is activated
     #tempSumPoint2 := #tempSumPoint2 - (#statUc2 / #statRthCool);
   END_IF;

   // Calculate Integrator 2
   #statUc2 := (#cycle * 0.5 * ((#tempSumPoint2 / #statCth2) + #statZInt2)) + #statUc2;
   #statZInt2 := #tempSumPoint2 / #statCth2;

   // Calculate Output Temperature
   #outTemp := #statUc2 + #ambTemp;
END_FUNCTION_BLOCK

